REGION Network 394
   RUNG wire#powerrail
      Contact( "EMS".Carrier[59].SDC_OUT.Faults.CarrierSpacingFault )
      Coil( "Carrier_59_Carrier_Spacing_Fault" )
   END_RUNG
   // the same network as SCL:
   "Carrier_59_Carrier_Spacing_Fault" := "EMS".Carrier[59].SDC_OUT.Faults.CarrierSpacingFault;
END_REGION

REGION Network 395
   RUNG wire#powerrail
      Move(in := "EMS".Carrier[60].SDC_OUT.Zone, out1 => "Carrier_60_Carrier_In_Zone")
   END_RUNG
   // the same network as SCL:
   "Carrier_60_Carrier_In_Zone" := "EMS".Carrier[60].SDC_OUT.Zone;
END_REGION

REGION Network 396
   RUNG wire#powerrail
      Move(in := "EMS".Carrier[60].SDC_OUT.CarrierNum, out1 => "Carrier_60_Carrier_Number_Echo")
   END_RUNG
   // the same network as SCL:
   "Carrier_60_Carrier_Number_Echo" := "EMS".Carrier[60].SDC_OUT.CarrierNum;
END_REGION

REGION Network 397
   RUNG wire#powerrail
      Move(in := "EMS".Carrier[60].SDC_OUT.CarrierPosition, out1 => "Carrier_60_Carrier_Position_Echo")
   END_RUNG
   // the same network as SCL:
   "Carrier_60_Carrier_Position_Echo" := "EMS".Carrier[60].SDC_OUT.CarrierPosition;
END_REGION

REGION Network 398
   RUNG wire#powerrail
      Move(in := "EMS".Carrier[60].SDC_OUT.NextCarrierNum, out1 => "Carrier_60_Next_Carrier_Number")
   END_RUNG
   // the same network as SCL:
   "Carrier_60_Next_Carrier_Number" := "EMS".Carrier[60].SDC_OUT.NextCarrierNum;
END_REGION

REGION Network 399
   RUNG wire#powerrail
      Move(in := "EMS".Carrier[60].SDC_OUT.NextStopPos, out1 => "Carrier_60_Next_Stop_Position")
   END_RUNG
   // the same network as SCL:
   "Carrier_60_Next_Stop_Position" := "EMS".Carrier[60].SDC_OUT.NextStopPos;
END_REGION

REGION Network 400
   RUNG wire#powerrail
      Move(in := "EMS".Carrier[60].SDC_OUT.DriveCmdSpeed, out1 => "Carrier_60_Drive_Command_Speed")
   END_RUNG
   // the same network as SCL:
   "Carrier_60_Drive_Command_Speed" := "EMS".Carrier[60].SDC_OUT.DriveCmdSpeed;
END_REGION

REGION Network 401
   RUNG wire#powerrail
      Move(in := "DuplicateCarrierNumber", out1 => "Carrier_60_Duplicate_Carrier_Number")
   END_RUNG
   // the same network as SCL:
   "Carrier_60_Duplicate_Carrier_Number" := "DuplicateCarrierNumber";
END_REGION

REGION Network 402
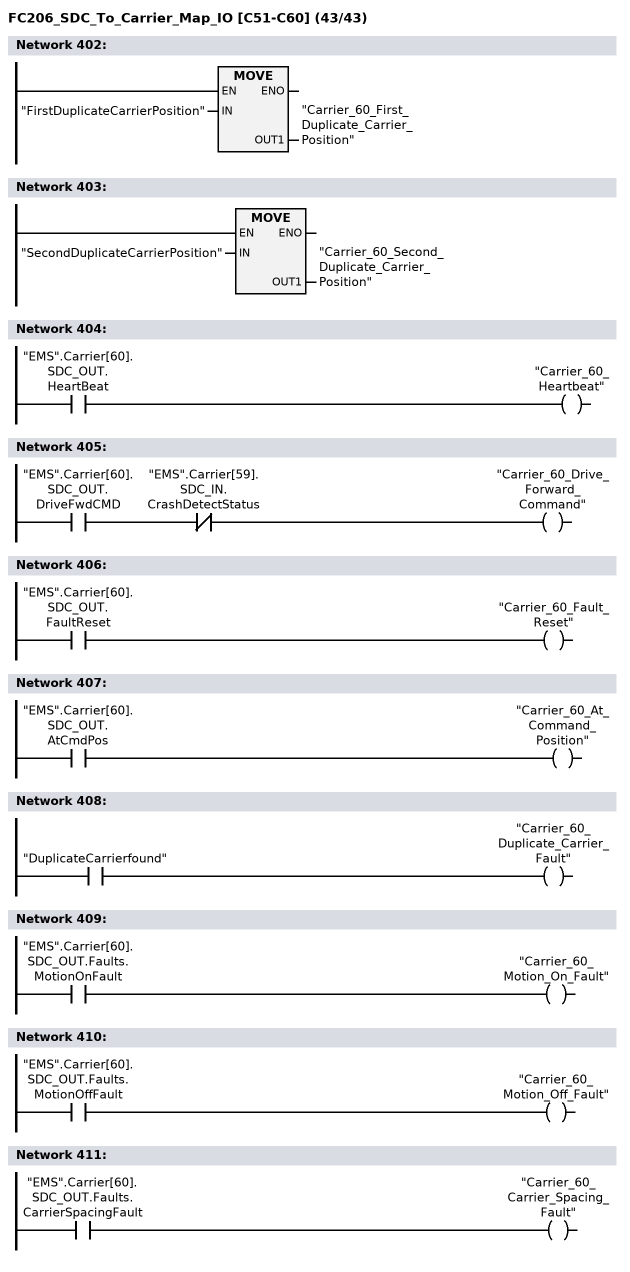
   RUNG wire#powerrail
      Move(in := "FirstDuplicateCarrierPosition", out1 => "Carrier_60_First_Duplicate_Carrier_Position")
   END_RUNG
   // the same network as SCL:
   "Carrier_60_First_Duplicate_Carrier_Position" := "FirstDuplicateCarrierPosition";
END_REGION

REGION Network 403
   RUNG wire#powerrail
      Move(in := "SecondDuplicateCarrierPosition", out1 => "Carrier_60_Second_Duplicate_Carrier_Position")
   END_RUNG
   // the same network as SCL:
   "Carrier_60_Second_Duplicate_Carrier_Position" := "SecondDuplicateCarrierPosition";
END_REGION

REGION Network 404
   RUNG wire#powerrail
      Contact( "EMS".Carrier[60].SDC_OUT.HeartBeat )
      Coil( "Carrier_60_Heartbeat" )
   END_RUNG
   // the same network as SCL:
   "Carrier_60_Heartbeat" := "EMS".Carrier[60].SDC_OUT.HeartBeat;
END_REGION

REGION Network 405
   RUNG wire#powerrail
      Contact( "EMS".Carrier[60].SDC_OUT.DriveFwdCMD )
      I_Contact( "EMS".Carrier[59].SDC_IN.CrashDetectStatus )
      Coil( "Carrier_60_Drive_Forward_Command" )
   END_RUNG
   // the same network as SCL:
   "Carrier_60_Drive_Forward_Command" := "EMS".Carrier[60].SDC_OUT.DriveFwdCMD AND NOT "EMS".Carrier[59].SDC_IN.CrashDetectStatus;
END_REGION

REGION Network 406
   RUNG wire#powerrail
      Contact( "EMS".Carrier[60].SDC_OUT.FaultReset )
      Coil( "Carrier_60_Fault_Reset" )
   END_RUNG
   // the same network as SCL:
   "Carrier_60_Fault_Reset" := "EMS".Carrier[60].SDC_OUT.FaultReset;
END_REGION

REGION Network 407
   RUNG wire#powerrail
      Contact( "EMS".Carrier[60].SDC_OUT.AtCmdPos )
      Coil( "Carrier_60_At_Command_Position" )
   END_RUNG
   // the same network as SCL:
   "Carrier_60_At_Command_Position" := "EMS".Carrier[60].SDC_OUT.AtCmdPos;
END_REGION

REGION Network 408
   RUNG wire#powerrail
      Contact( "DuplicateCarrierfound" )
      Coil( "Carrier_60_Duplicate_Carrier_Fault" )
   END_RUNG
   // the same network as SCL:
   "Carrier_60_Duplicate_Carrier_Fault" := "DuplicateCarrierfound";
END_REGION

REGION Network 409
   RUNG wire#powerrail
      Contact( "EMS".Carrier[60].SDC_OUT.Faults.MotionOnFault )
      Coil( "Carrier_60_Motion_On_Fault" )
   END_RUNG
   // the same network as SCL:
   "Carrier_60_Motion_On_Fault" := "EMS".Carrier[60].SDC_OUT.Faults.MotionOnFault;
END_REGION

REGION Network 410
   RUNG wire#powerrail
      Contact( "EMS".Carrier[60].SDC_OUT.Faults.MotionOffFault )
      Coil( "Carrier_60_Motion_Off_Fault" )
   END_RUNG
   // the same network as SCL:
   "Carrier_60_Motion_Off_Fault" := "EMS".Carrier[60].SDC_OUT.Faults.MotionOffFault;
END_REGION

REGION Network 411
   RUNG wire#powerrail
      Contact( "EMS".Carrier[60].SDC_OUT.Faults.CarrierSpacingFault )
      Coil( "Carrier_60_Carrier_Spacing_Fault" )
   END_RUNG
   // the same network as SCL:
   "Carrier_60_Carrier_Spacing_Fault" := "EMS".Carrier[60].SDC_OUT.Faults.CarrierSpacingFault;
END_REGION
END_FUNCTION

FUNCTION "FC207_SDC_To_Carrier_Map_IO [C61-C70]" : Void   // FC207, LAD
{ S7_Optimized_Access := 'TRUE' }
VERSION : 0.1
BEGIN

REGION Network 1
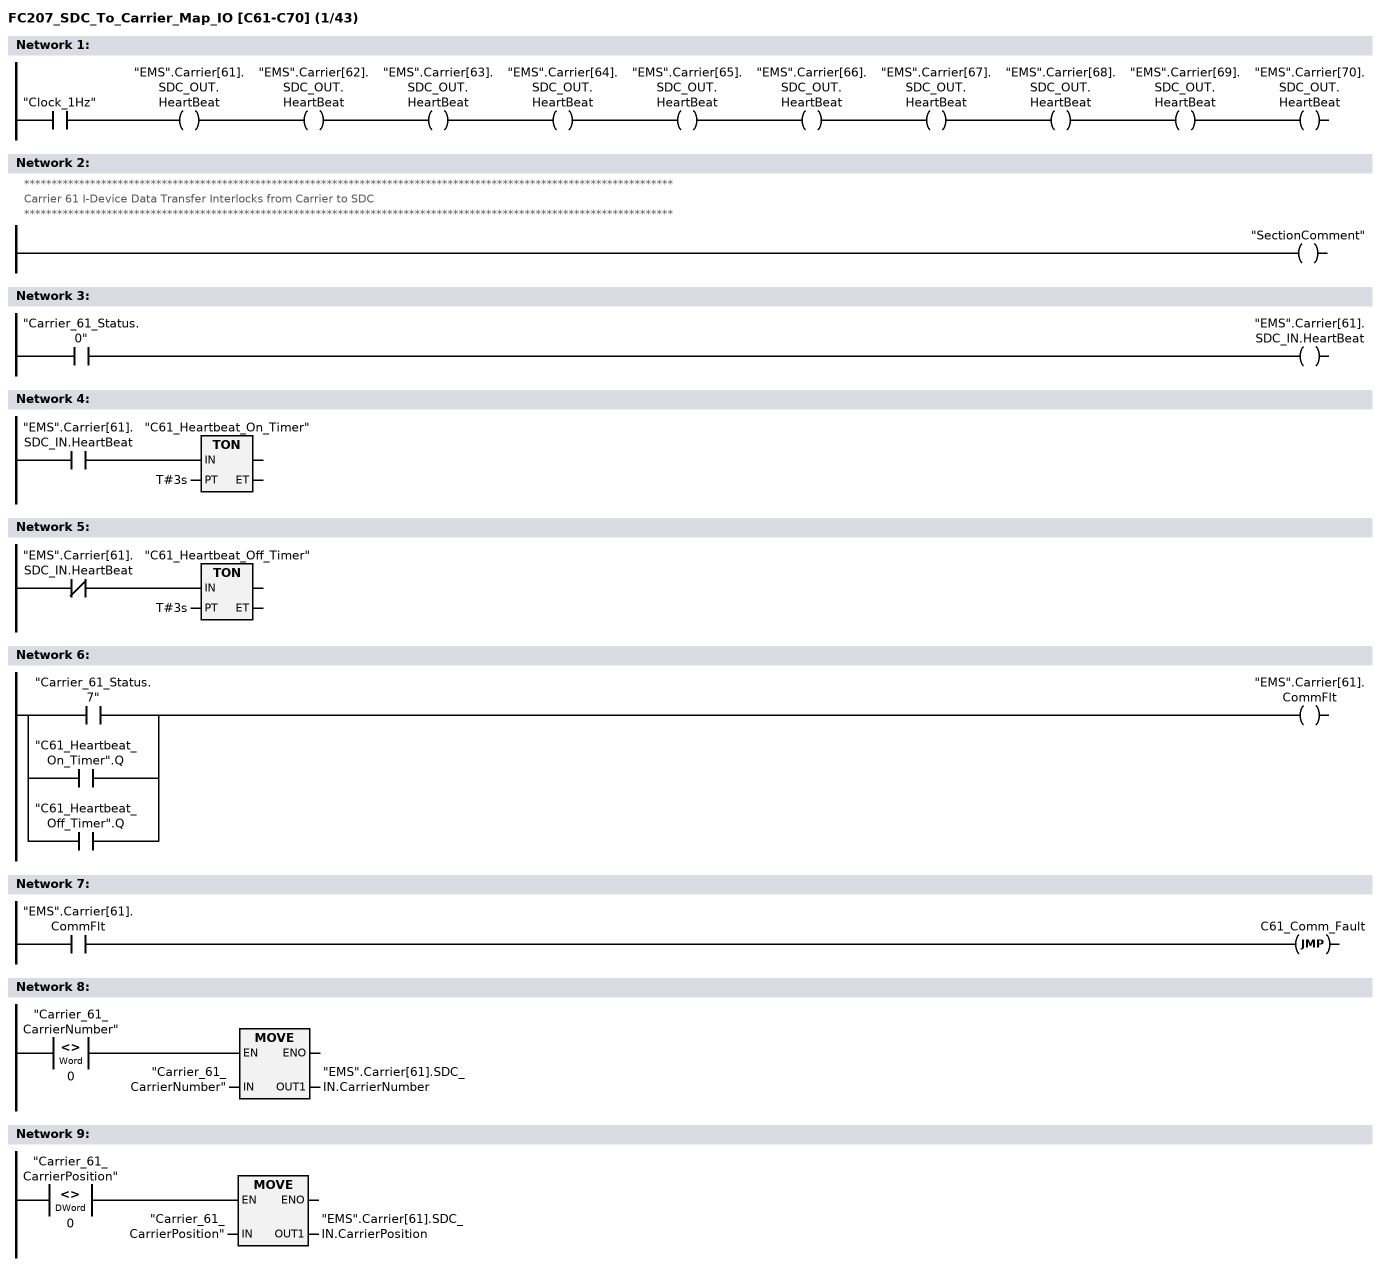
   RUNG wire#powerrail
      Contact( "Clock_1Hz" )
      Coil( "EMS".Carrier[61].SDC_OUT.HeartBeat )
      Coil( "EMS".Carrier[62].SDC_OUT.HeartBeat )
      Coil( "EMS".Carrier[63].SDC_OUT.HeartBeat )
      Coil( "EMS".Carrier[64].SDC_OUT.HeartBeat )
      Coil( "EMS".Carrier[65].SDC_OUT.HeartBeat )
      Coil( "EMS".Carrier[66].SDC_OUT.HeartBeat )
      Coil( "EMS".Carrier[67].SDC_OUT.HeartBeat )
      Coil( "EMS".Carrier[68].SDC_OUT.HeartBeat )
      Coil( "EMS".Carrier[69].SDC_OUT.HeartBeat )
      Coil( "EMS".Carrier[70].SDC_OUT.HeartBeat )
   END_RUNG
   // the same network as SCL:
   "EMS".Carrier[61].SDC_OUT.HeartBeat := "Clock_1Hz";
   "EMS".Carrier[62].SDC_OUT.HeartBeat := "Clock_1Hz";
   "EMS".Carrier[63].SDC_OUT.HeartBeat := "Clock_1Hz";
   "EMS".Carrier[64].SDC_OUT.HeartBeat := "Clock_1Hz";
   "EMS".Carrier[65].SDC_OUT.HeartBeat := "Clock_1Hz";
   "EMS".Carrier[66].SDC_OUT.HeartBeat := "Clock_1Hz";
   "EMS".Carrier[67].SDC_OUT.HeartBeat := "Clock_1Hz";
   "EMS".Carrier[68].SDC_OUT.HeartBeat := "Clock_1Hz";
   "EMS".Carrier[69].SDC_OUT.HeartBeat := "Clock_1Hz";
   "EMS".Carrier[70].SDC_OUT.HeartBeat := "Clock_1Hz";
END_REGION

REGION Network 2
   // **********************************************************************************************************************
   // 
   // Carrier 61 I-Device Data Transfer Interlocks from Carrier to SDC
   // 
   // **********************************************************************************************************************
   RUNG wire#powerrail
      Coil( "SectionComment" )
   END_RUNG
   // the same network as SCL:
   "SectionComment" := TRUE;
END_REGION

REGION Network 3
   RUNG wire#powerrail
      Contact( "Carrier_61_Status.0" )
      Coil( "EMS".Carrier[61].SDC_IN.HeartBeat )
   END_RUNG
   // the same network as SCL:
   "EMS".Carrier[61].SDC_IN.HeartBeat := "Carrier_61_Status.0";
END_REGION

REGION Network 4
   "C61_Heartbeat_On_Timer".TON(IN := "EMS".Carrier[61].SDC_IN.HeartBeat, PT := T#3s);
END_REGION

REGION Network 5
   "C61_Heartbeat_Off_Timer".TON(IN := NOT "EMS".Carrier[61].SDC_IN.HeartBeat, PT := T#3s);
END_REGION

REGION Network 6
   RUNG wire#powerrail
      Contact( "Carrier_61_Status.7" )
      wire#w1
      Coil( "EMS".Carrier[61].CommFlt )
   END_RUNG
   RUNG wire#powerrail
      Contact( "C61_Heartbeat_On_Timer".Q )
   END_RUNG wire#w1
   RUNG wire#powerrail
      Contact( "C61_Heartbeat_Off_Timer".Q )
   END_RUNG wire#w1
   // the same network as SCL:
   "EMS".Carrier[61].CommFlt := "Carrier_61_Status.7" OR "C61_Heartbeat_On_Timer".Q OR "C61_Heartbeat_Off_Timer".Q;
END_REGION

REGION Network 7
   RUNG wire#powerrail
      Contact( "EMS".Carrier[61].CommFlt )
      JumpCoil( C61_Comm_Fault )
   END_RUNG
   // the same network as SCL:
   IF "EMS".Carrier[61].CommFlt THEN GOTO C61_Comm_Fault; END_IF;
END_REGION

REGION Network 8
   RUNG wire#powerrail
      { S7_Templates := "SrcType := Word" } NE_Contact(in1 := "Carrier_61_CarrierNumber", in2 := 0)
      Move(in := "Carrier_61_CarrierNumber", out1 => "EMS".Carrier[61].SDC_IN.CarrierNumber)
   END_RUNG
   // the same network as SCL:
   IF "Carrier_61_CarrierNumber" <> 0 THEN
       "EMS".Carrier[61].SDC_IN.CarrierNumber := "Carrier_61_CarrierNumber";
   END_IF;
END_REGION

REGION Network 9
   RUNG wire#powerrail
      { S7_Templates := "SrcType := DWord" } NE_Contact(in1 := "Carrier_61_CarrierPosition", in2 := 0)
      Move(in := "Carrier_61_CarrierPosition", out1 => "EMS".Carrier[61].SDC_IN.CarrierPosition)
   END_RUNG
   // the same network as SCL:
   IF "Carrier_61_CarrierPosition" <> 0 THEN
       "EMS".Carrier[61].SDC_IN.CarrierPosition := "Carrier_61_CarrierPosition";
   END_IF;
END_REGION

REGION Network 10
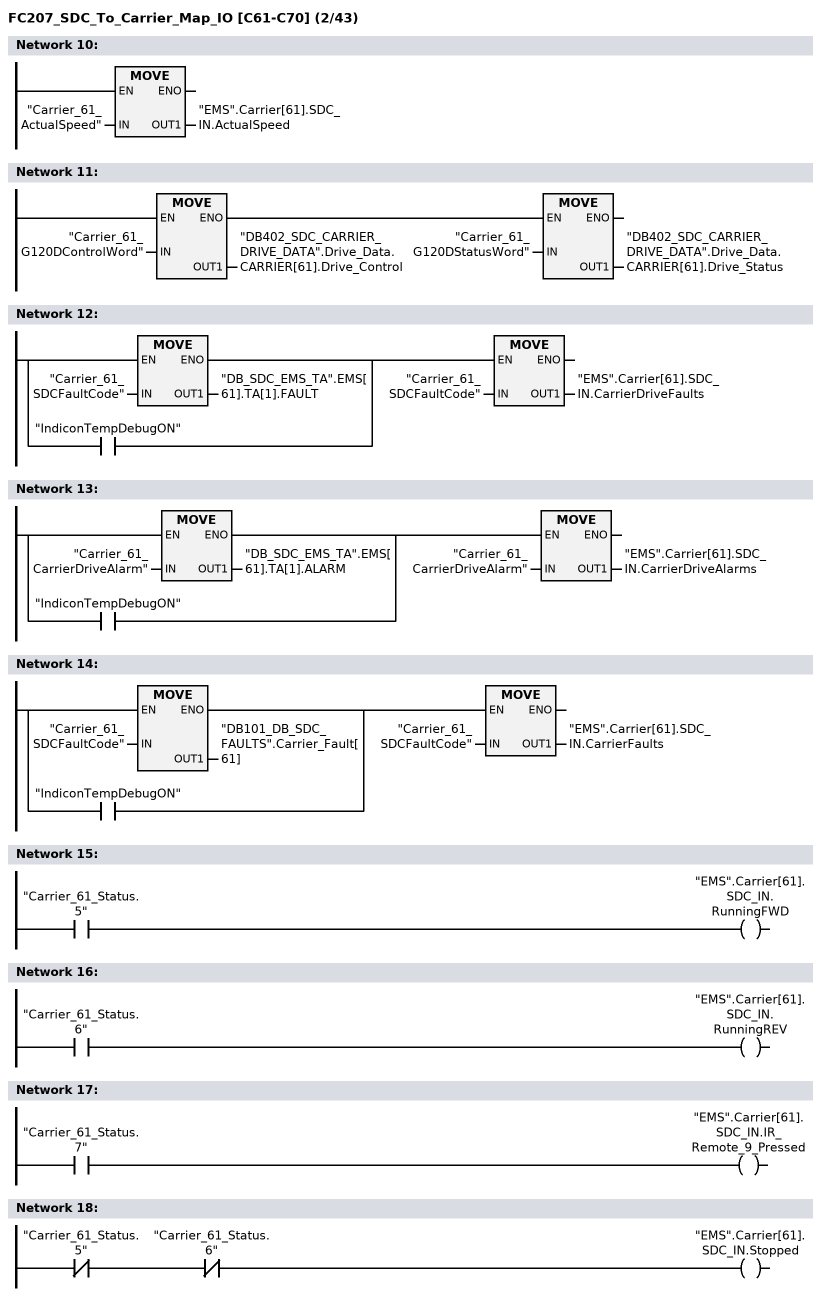
   RUNG wire#powerrail
      Move(in := "Carrier_61_ActualSpeed", out1 => "EMS".Carrier[61].SDC_IN.ActualSpeed)
   END_RUNG
   // the same network as SCL:
   "EMS".Carrier[61].SDC_IN.ActualSpeed := "Carrier_61_ActualSpeed";
END_REGION

REGION Network 11
   RUNG wire#powerrail
      Move(in := "Carrier_61_G120DControlWord", out1 => "DB402_SDC_CARRIER_DRIVE_DATA".Drive_Data.CARRIER[61].Drive_Control)
      Move(in := "Carrier_61_G120DStatusWord", out1 => "DB402_SDC_CARRIER_DRIVE_DATA".Drive_Data.CARRIER[61].Drive_Status)
   END_RUNG
   // the same network as SCL:
   "DB402_SDC_CARRIER_DRIVE_DATA".Drive_Data.CARRIER[61].Drive_Control := "Carrier_61_G120DControlWord";
   "DB402_SDC_CARRIER_DRIVE_DATA".Drive_Data.CARRIER[61].Drive_Status := "Carrier_61_G120DStatusWord";
END_REGION

REGION Network 12
   RUNG wire#powerrail
      Move(in := "Carrier_61_SDCFaultCode", out1 => "DB_SDC_EMS_TA".EMS[61].TA[1].FAULT)
      wire#w1
      Move(in := "Carrier_61_SDCFaultCode", out1 => "EMS".Carrier[61].SDC_IN.CarrierDriveFaults)
   END_RUNG
   RUNG wire#powerrail
      Contact( "IndiconTempDebugON" )
   END_RUNG wire#w1
   // the same network as SCL:
   "DB_SDC_EMS_TA".EMS[61].TA[1].FAULT := "Carrier_61_SDCFaultCode";
   IF TRUE OR "IndiconTempDebugON" THEN
       "EMS".Carrier[61].SDC_IN.CarrierDriveFaults := "Carrier_61_SDCFaultCode";
   END_IF;
END_REGION

REGION Network 13
   RUNG wire#powerrail
      Move(in := "Carrier_61_CarrierDriveAlarm", out1 => "DB_SDC_EMS_TA".EMS[61].TA[1].ALARM)
      wire#w1
      Move(in := "Carrier_61_CarrierDriveAlarm", out1 => "EMS".Carrier[61].SDC_IN.CarrierDriveAlarms)
   END_RUNG
   RUNG wire#powerrail
      Contact( "IndiconTempDebugON" )
   END_RUNG wire#w1
   // the same network as SCL:
   "DB_SDC_EMS_TA".EMS[61].TA[1].ALARM := "Carrier_61_CarrierDriveAlarm";
   IF TRUE OR "IndiconTempDebugON" THEN
       "EMS".Carrier[61].SDC_IN.CarrierDriveAlarms := "Carrier_61_CarrierDriveAlarm";
   END_IF;
END_REGION

REGION Network 14
   RUNG wire#powerrail
      Move(in := "Carrier_61_SDCFaultCode", out1 => "DB101_DB_SDC_FAULTS".Carrier_Fault[61])
      wire#w1
      Move(in := "Carrier_61_SDCFaultCode", out1 => "EMS".Carrier[61].SDC_IN.CarrierFaults)
   END_RUNG
   RUNG wire#powerrail
      Contact( "IndiconTempDebugON" )
   END_RUNG wire#w1
   // the same network as SCL:
   "DB101_DB_SDC_FAULTS".Carrier_Fault[61] := "Carrier_61_SDCFaultCode";
   IF TRUE OR "IndiconTempDebugON" THEN
       "EMS".Carrier[61].SDC_IN.CarrierFaults := "Carrier_61_SDCFaultCode";
   END_IF;
END_REGION

REGION Network 15
   RUNG wire#powerrail
      Contact( "Carrier_61_Status.5" )
      Coil( "EMS".Carrier[61].SDC_IN.RunningFWD )
   END_RUNG
   // the same network as SCL:
   "EMS".Carrier[61].SDC_IN.RunningFWD := "Carrier_61_Status.5";
END_REGION

REGION Network 16
   RUNG wire#powerrail
      Contact( "Carrier_61_Status.6" )
      Coil( "EMS".Carrier[61].SDC_IN.RunningREV )
   END_RUNG
   // the same network as SCL:
   "EMS".Carrier[61].SDC_IN.RunningREV := "Carrier_61_Status.6";
END_REGION

REGION Network 17
   RUNG wire#powerrail
      Contact( "Carrier_61_Status.7" )
      Coil( "EMS".Carrier[61].SDC_IN.IR_Remote_9_Pressed )
   END_RUNG
   // the same network as SCL:
   "EMS".Carrier[61].SDC_IN.IR_Remote_9_Pressed := "Carrier_61_Status.7";
END_REGION

REGION Network 18
   RUNG wire#powerrail
      I_Contact( "Carrier_61_Status.5" )
      I_Contact( "Carrier_61_Status.6" )
      Coil( "EMS".Carrier[61].SDC_IN.Stopped )
   END_RUNG
   // the same network as SCL:
   "EMS".Carrier[61].SDC_IN.Stopped := NOT "Carrier_61_Status.5" AND NOT "Carrier_61_Status.6";
END_REGION

REGION Network 19
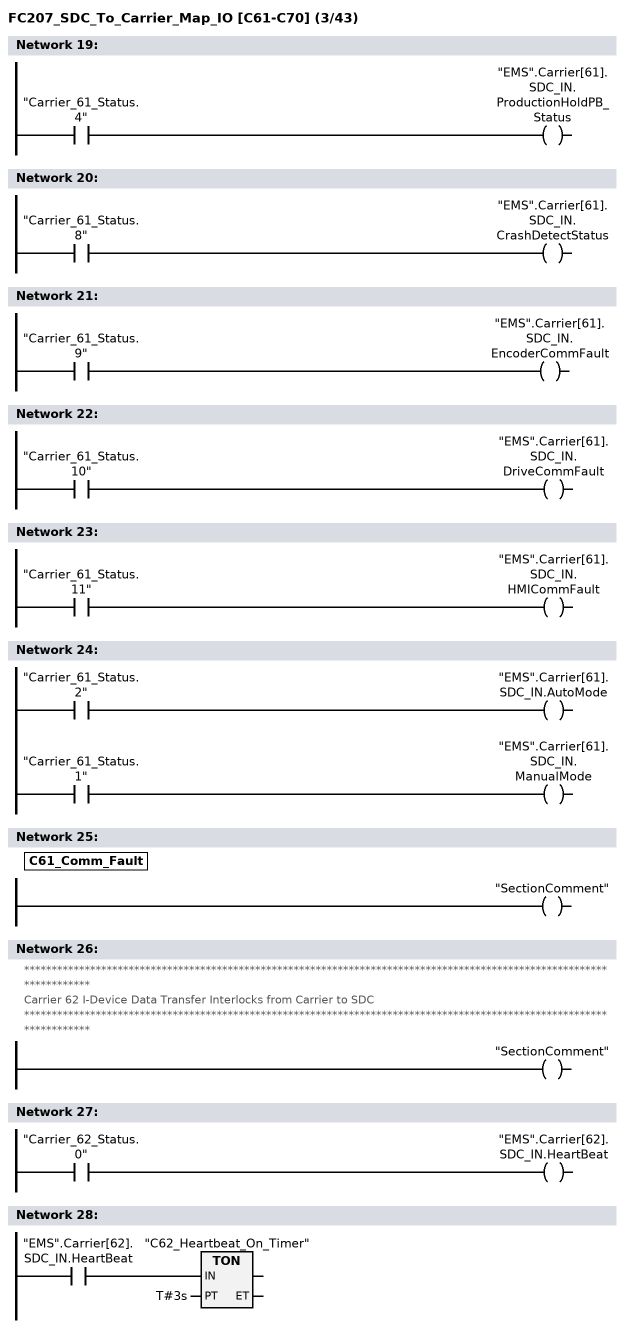
   RUNG wire#powerrail
      Contact( "Carrier_61_Status.4" )
      Coil( "EMS".Carrier[61].SDC_IN.ProductionHoldPB_Status )
   END_RUNG
   // the same network as SCL:
   "EMS".Carrier[61].SDC_IN.ProductionHoldPB_Status := "Carrier_61_Status.4";
END_REGION

REGION Network 20
   RUNG wire#powerrail
      Contact( "Carrier_61_Status.8" )
      Coil( "EMS".Carrier[61].SDC_IN.CrashDetectStatus )
   END_RUNG
   // the same network as SCL:
   "EMS".Carrier[61].SDC_IN.CrashDetectStatus := "Carrier_61_Status.8";
END_REGION

REGION Network 21
   RUNG wire#powerrail
      Contact( "Carrier_61_Status.9" )
      Coil( "EMS".Carrier[61].SDC_IN.EncoderCommFault )
   END_RUNG
   // the same network as SCL:
   "EMS".Carrier[61].SDC_IN.EncoderCommFault := "Carrier_61_Status.9";
END_REGION

REGION Network 22
   RUNG wire#powerrail
      Contact( "Carrier_61_Status.10" )
      Coil( "EMS".Carrier[61].SDC_IN.DriveCommFault )
   END_RUNG
   // the same network as SCL:
   "EMS".Carrier[61].SDC_IN.DriveCommFault := "Carrier_61_Status.10";
END_REGION

REGION Network 23
   RUNG wire#powerrail
      Contact( "Carrier_61_Status.11" )
      Coil( "EMS".Carrier[61].SDC_IN.HMICommFault )
   END_RUNG
   // the same network as SCL:
   "EMS".Carrier[61].SDC_IN.HMICommFault := "Carrier_61_Status.11";
END_REGION

REGION Network 24
   RUNG wire#powerrail
      Contact( "Carrier_61_Status.2" )
      Coil( "EMS".Carrier[61].SDC_IN.AutoMode )
   END_RUNG
   RUNG wire#powerrail
      Contact( "Carrier_61_Status.1" )
      Coil( "EMS".Carrier[61].SDC_IN.ManualMode )
   END_RUNG
   // the same network as SCL:
   "EMS".Carrier[61].SDC_IN.AutoMode := "Carrier_61_Status.2";
   "EMS".Carrier[61].SDC_IN.ManualMode := "Carrier_61_Status.1";
END_REGION

REGION Network 25
   Label( C61_Comm_Fault )
   RUNG wire#powerrail
      Coil( "SectionComment" )
   END_RUNG
   // the same network as SCL:
   C61_Comm_Fault:
   "SectionComment" := TRUE;
END_REGION

REGION Network 26
   // **********************************************************************************************************************
   // 
   // Carrier 62 I-Device Data Transfer Interlocks from Carrier to SDC
   // 
   // **********************************************************************************************************************
   RUNG wire#powerrail
      Coil( "SectionComment" )
   END_RUNG
   // the same network as SCL:
   "SectionComment" := TRUE;
END_REGION

REGION Network 27
   RUNG wire#powerrail
      Contact( "Carrier_62_Status.0" )
      Coil( "EMS".Carrier[62].SDC_IN.HeartBeat )
   END_RUNG
   // the same network as SCL:
   "EMS".Carrier[62].SDC_IN.HeartBeat := "Carrier_62_Status.0";
END_REGION

REGION Network 28
   "C62_Heartbeat_On_Timer".TON(IN := "EMS".Carrier[62].SDC_IN.HeartBeat, PT := T#3s);
END_REGION

REGION Network 29
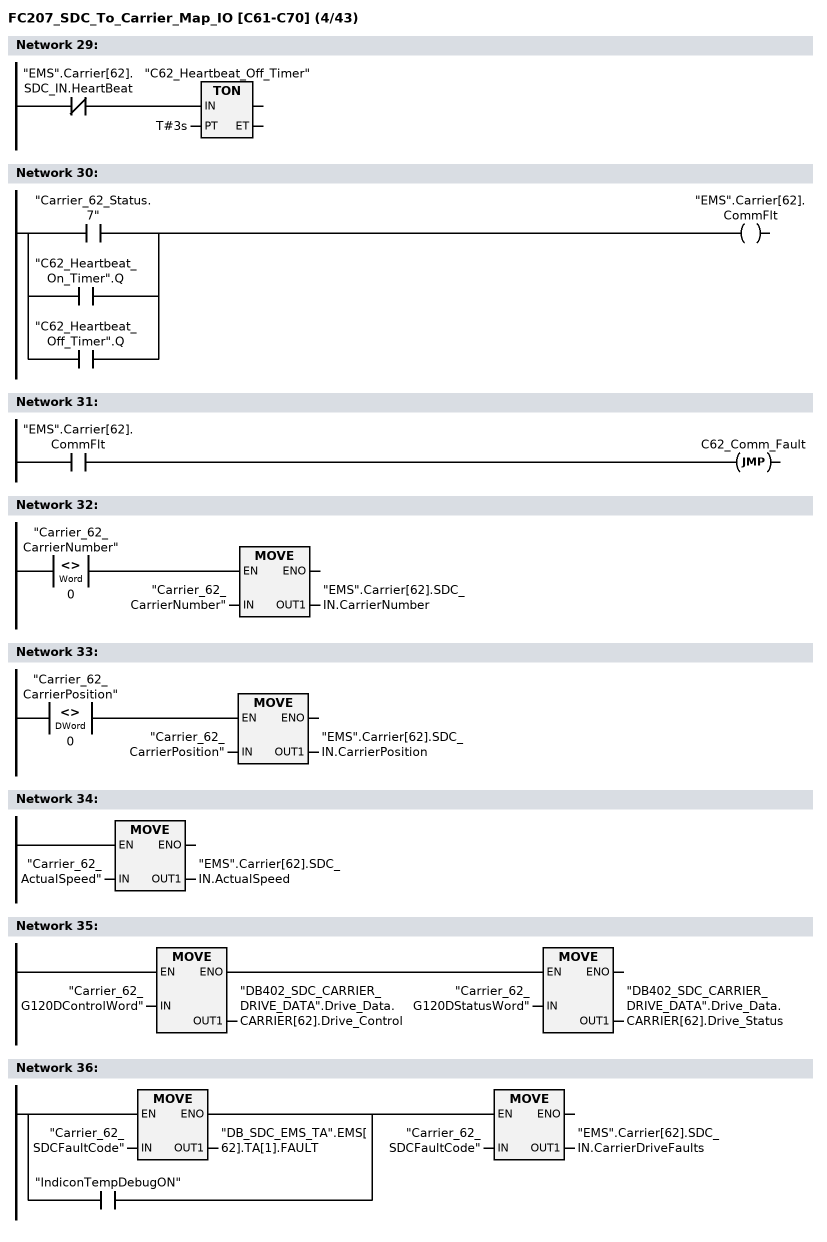
   "C62_Heartbeat_Off_Timer".TON(IN := NOT "EMS".Carrier[62].SDC_IN.HeartBeat, PT := T#3s);
END_REGION

REGION Network 30
   RUNG wire#powerrail
      Contact( "Carrier_62_Status.7" )
      wire#w1
      Coil( "EMS".Carrier[62].CommFlt )
   END_RUNG
   RUNG wire#powerrail
      Contact( "C62_Heartbeat_On_Timer".Q )
   END_RUNG wire#w1
   RUNG wire#powerrail
      Contact( "C62_Heartbeat_Off_Timer".Q )
   END_RUNG wire#w1
   // the same network as SCL:
   "EMS".Carrier[62].CommFlt := "Carrier_62_Status.7" OR "C62_Heartbeat_On_Timer".Q OR "C62_Heartbeat_Off_Timer".Q;
END_REGION

REGION Network 31
   RUNG wire#powerrail
      Contact( "EMS".Carrier[62].CommFlt )
      JumpCoil( C62_Comm_Fault )
   END_RUNG
   // the same network as SCL:
   IF "EMS".Carrier[62].CommFlt THEN GOTO C62_Comm_Fault; END_IF;
END_REGION

REGION Network 32
   RUNG wire#powerrail
      { S7_Templates := "SrcType := Word" } NE_Contact(in1 := "Carrier_62_CarrierNumber", in2 := 0)
      Move(in := "Carrier_62_CarrierNumber", out1 => "EMS".Carrier[62].SDC_IN.CarrierNumber)
   END_RUNG
   // the same network as SCL:
   IF "Carrier_62_CarrierNumber" <> 0 THEN
       "EMS".Carrier[62].SDC_IN.CarrierNumber := "Carrier_62_CarrierNumber";
   END_IF;
END_REGION

REGION Network 33
   RUNG wire#powerrail
      { S7_Templates := "SrcType := DWord" } NE_Contact(in1 := "Carrier_62_CarrierPosition", in2 := 0)
      Move(in := "Carrier_62_CarrierPosition", out1 => "EMS".Carrier[62].SDC_IN.CarrierPosition)
   END_RUNG
   // the same network as SCL:
   IF "Carrier_62_CarrierPosition" <> 0 THEN
       "EMS".Carrier[62].SDC_IN.CarrierPosition := "Carrier_62_CarrierPosition";
   END_IF;
END_REGION

REGION Network 34
   RUNG wire#powerrail
      Move(in := "Carrier_62_ActualSpeed", out1 => "EMS".Carrier[62].SDC_IN.ActualSpeed)
   END_RUNG
   // the same network as SCL:
   "EMS".Carrier[62].SDC_IN.ActualSpeed := "Carrier_62_ActualSpeed";
END_REGION

REGION Network 35
   RUNG wire#powerrail
      Move(in := "Carrier_62_G120DControlWord", out1 => "DB402_SDC_CARRIER_DRIVE_DATA".Drive_Data.CARRIER[62].Drive_Control)
      Move(in := "Carrier_62_G120DStatusWord", out1 => "DB402_SDC_CARRIER_DRIVE_DATA".Drive_Data.CARRIER[62].Drive_Status)
   END_RUNG
   // the same network as SCL:
   "DB402_SDC_CARRIER_DRIVE_DATA".Drive_Data.CARRIER[62].Drive_Control := "Carrier_62_G120DControlWord";
   "DB402_SDC_CARRIER_DRIVE_DATA".Drive_Data.CARRIER[62].Drive_Status := "Carrier_62_G120DStatusWord";
END_REGION

REGION Network 36
   RUNG wire#powerrail
      Move(in := "Carrier_62_SDCFaultCode", out1 => "DB_SDC_EMS_TA".EMS[62].TA[1].FAULT)
      wire#w1
      Move(in := "Carrier_62_SDCFaultCode", out1 => "EMS".Carrier[62].SDC_IN.CarrierDriveFaults)
   END_RUNG
   RUNG wire#powerrail
      Contact( "IndiconTempDebugON" )
   END_RUNG wire#w1
   // the same network as SCL:
   "DB_SDC_EMS_TA".EMS[62].TA[1].FAULT := "Carrier_62_SDCFaultCode";
   IF TRUE OR "IndiconTempDebugON" THEN
       "EMS".Carrier[62].SDC_IN.CarrierDriveFaults := "Carrier_62_SDCFaultCode";
   END_IF;
END_REGION

REGION Network 37
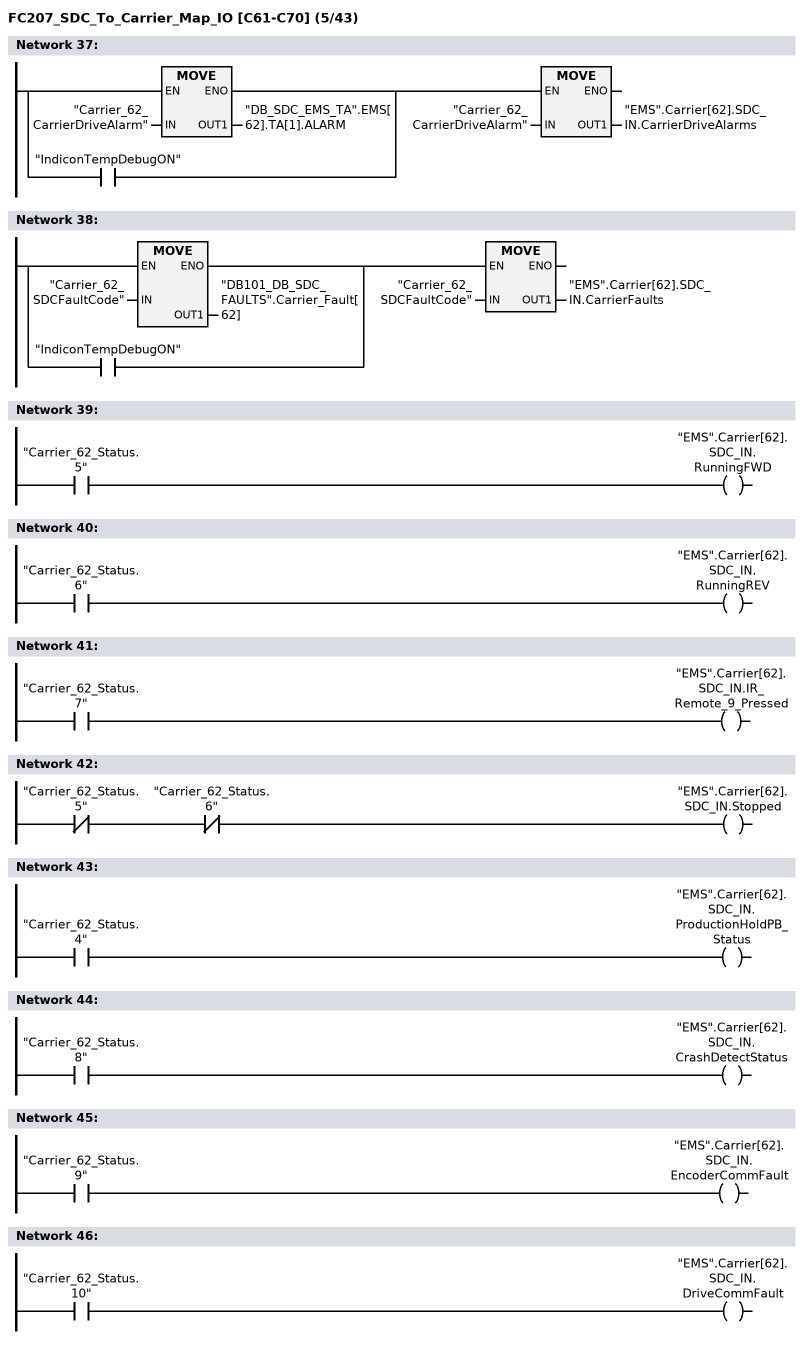
   RUNG wire#powerrail
      Move(in := "Carrier_62_CarrierDriveAlarm", out1 => "DB_SDC_EMS_TA".EMS[62].TA[1].ALARM)
      wire#w1
      Move(in := "Carrier_62_CarrierDriveAlarm", out1 => "EMS".Carrier[62].SDC_IN.CarrierDriveAlarms)
   END_RUNG
   RUNG wire#powerrail
      Contact( "IndiconTempDebugON" )
   END_RUNG wire#w1
   // the same network as SCL:
   "DB_SDC_EMS_TA".EMS[62].TA[1].ALARM := "Carrier_62_CarrierDriveAlarm";
   IF TRUE OR "IndiconTempDebugON" THEN
       "EMS".Carrier[62].SDC_IN.CarrierDriveAlarms := "Carrier_62_CarrierDriveAlarm";
   END_IF;
END_REGION

REGION Network 38
   RUNG wire#powerrail
      Move(in := "Carrier_62_SDCFaultCode", out1 => "DB101_DB_SDC_FAULTS".Carrier_Fault[62])
      wire#w1
      Move(in := "Carrier_62_SDCFaultCode", out1 => "EMS".Carrier[62].SDC_IN.CarrierFaults)
   END_RUNG
   RUNG wire#powerrail
      Contact( "IndiconTempDebugON" )
   END_RUNG wire#w1
   // the same network as SCL:
   "DB101_DB_SDC_FAULTS".Carrier_Fault[62] := "Carrier_62_SDCFaultCode";
   IF TRUE OR "IndiconTempDebugON" THEN
       "EMS".Carrier[62].SDC_IN.CarrierFaults := "Carrier_62_SDCFaultCode";
   END_IF;
END_REGION

REGION Network 39
   RUNG wire#powerrail
      Contact( "Carrier_62_Status.5" )
      Coil( "EMS".Carrier[62].SDC_IN.RunningFWD )
   END_RUNG
   // the same network as SCL:
   "EMS".Carrier[62].SDC_IN.RunningFWD := "Carrier_62_Status.5";
END_REGION

REGION Network 40
   RUNG wire#powerrail
      Contact( "Carrier_62_Status.6" )
      Coil( "EMS".Carrier[62].SDC_IN.RunningREV )
   END_RUNG
   // the same network as SCL:
   "EMS".Carrier[62].SDC_IN.RunningREV := "Carrier_62_Status.6";
END_REGION

REGION Network 41
   RUNG wire#powerrail
      Contact( "Carrier_62_Status.7" )
      Coil( "EMS".Carrier[62].SDC_IN.IR_Remote_9_Pressed )
   END_RUNG
   // the same network as SCL:
   "EMS".Carrier[62].SDC_IN.IR_Remote_9_Pressed := "Carrier_62_Status.7";
END_REGION

REGION Network 42
   RUNG wire#powerrail
      I_Contact( "Carrier_62_Status.5" )
      I_Contact( "Carrier_62_Status.6" )
      Coil( "EMS".Carrier[62].SDC_IN.Stopped )
   END_RUNG
   // the same network as SCL:
   "EMS".Carrier[62].SDC_IN.Stopped := NOT "Carrier_62_Status.5" AND NOT "Carrier_62_Status.6";
END_REGION

REGION Network 43
   RUNG wire#powerrail
      Contact( "Carrier_62_Status.4" )
      Coil( "EMS".Carrier[62].SDC_IN.ProductionHoldPB_Status )
   END_RUNG
   // the same network as SCL:
   "EMS".Carrier[62].SDC_IN.ProductionHoldPB_Status := "Carrier_62_Status.4";
END_REGION

REGION Network 44
   RUNG wire#powerrail
      Contact( "Carrier_62_Status.8" )
      Coil( "EMS".Carrier[62].SDC_IN.CrashDetectStatus )
   END_RUNG
   // the same network as SCL:
   "EMS".Carrier[62].SDC_IN.CrashDetectStatus := "Carrier_62_Status.8";
END_REGION

REGION Network 45
   RUNG wire#powerrail
      Contact( "Carrier_62_Status.9" )
      Coil( "EMS".Carrier[62].SDC_IN.EncoderCommFault )
   END_RUNG
   // the same network as SCL:
   "EMS".Carrier[62].SDC_IN.EncoderCommFault := "Carrier_62_Status.9";
END_REGION

REGION Network 46
   RUNG wire#powerrail
      Contact( "Carrier_62_Status.10" )
      Coil( "EMS".Carrier[62].SDC_IN.DriveCommFault )
   END_RUNG
   // the same network as SCL:
   "EMS".Carrier[62].SDC_IN.DriveCommFault := "Carrier_62_Status.10";
END_REGION

REGION Network 47
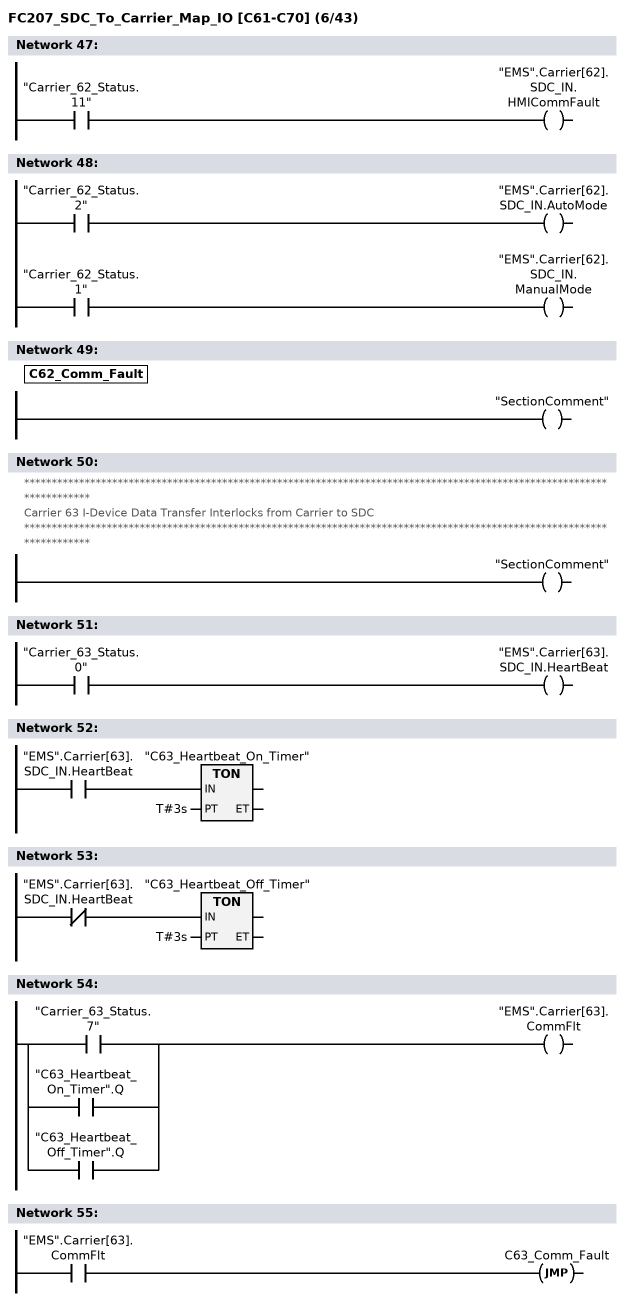
   RUNG wire#powerrail
      Contact( "Carrier_62_Status.11" )
      Coil( "EMS".Carrier[62].SDC_IN.HMICommFault )
   END_RUNG
   // the same network as SCL:
   "EMS".Carrier[62].SDC_IN.HMICommFault := "Carrier_62_Status.11";
END_REGION

REGION Network 48
   RUNG wire#powerrail
      Contact( "Carrier_62_Status.2" )
      Coil( "EMS".Carrier[62].SDC_IN.AutoMode )
   END_RUNG
   RUNG wire#powerrail
      Contact( "Carrier_62_Status.1" )
      Coil( "EMS".Carrier[62].SDC_IN.ManualMode )
   END_RUNG
   // the same network as SCL:
   "EMS".Carrier[62].SDC_IN.AutoMode := "Carrier_62_Status.2";
   "EMS".Carrier[62].SDC_IN.ManualMode := "Carrier_62_Status.1";
END_REGION

REGION Network 49
   Label( C62_Comm_Fault )
   RUNG wire#powerrail
      Coil( "SectionComment" )
   END_RUNG
   // the same network as SCL:
   C62_Comm_Fault:
   "SectionComment" := TRUE;
END_REGION

REGION Network 50
   // **********************************************************************************************************************
   // 
   // Carrier 63 I-Device Data Transfer Interlocks from Carrier to SDC
   // 
   // **********************************************************************************************************************
   RUNG wire#powerrail
      Coil( "SectionComment" )
   END_RUNG
   // the same network as SCL:
   "SectionComment" := TRUE;
END_REGION

REGION Network 51
   RUNG wire#powerrail
      Contact( "Carrier_63_Status.0" )
      Coil( "EMS".Carrier[63].SDC_IN.HeartBeat )
   END_RUNG
   // the same network as SCL:
   "EMS".Carrier[63].SDC_IN.HeartBeat := "Carrier_63_Status.0";
END_REGION

REGION Network 52
   "C63_Heartbeat_On_Timer".TON(IN := "EMS".Carrier[63].SDC_IN.HeartBeat, PT := T#3s);
END_REGION

REGION Network 53
   "C63_Heartbeat_Off_Timer".TON(IN := NOT "EMS".Carrier[63].SDC_IN.HeartBeat, PT := T#3s);
END_REGION

REGION Network 54
   RUNG wire#powerrail
      Contact( "Carrier_63_Status.7" )
      wire#w1
      Coil( "EMS".Carrier[63].CommFlt )
   END_RUNG
   RUNG wire#powerrail
      Contact( "C63_Heartbeat_On_Timer".Q )
   END_RUNG wire#w1
   RUNG wire#powerrail
      Contact( "C63_Heartbeat_Off_Timer".Q )
   END_RUNG wire#w1
   // the same network as SCL:
   "EMS".Carrier[63].CommFlt := "Carrier_63_Status.7" OR "C63_Heartbeat_On_Timer".Q OR "C63_Heartbeat_Off_Timer".Q;
END_REGION

REGION Network 55
   RUNG wire#powerrail
      Contact( "EMS".Carrier[63].CommFlt )
      JumpCoil( C63_Comm_Fault )
   END_RUNG
   // the same network as SCL:
   IF "EMS".Carrier[63].CommFlt THEN GOTO C63_Comm_Fault; END_IF;
END_REGION

REGION Network 56
